// TIA Portal project "Lagerbereich_0" (V20)

(* hardware
DEVICE "S7-1500/ET200MP-Station_1"  S7-1500 station
   slot 0: "Profilschiene_0"  Rack  6ES7 590-1***0-0AA0
   slot 1: "PLC_1"  CPU 1513-1 PN  6ES7 513-1AM03-0AB0  V4.0
      slot 3: "CPU-Display_1"  6ES7591-1AA00-0AA0
      slot 32768: "PROFINET-Schnittstelle_1"  X1
         slot 32769: "Port_1"  X1 P1
         slot 32770: "Port_2"  X1 P2
      slot 34817: "Virtual CP interface port_1"  Virtual CP interface port  Virtual CP interface port FW V4.0
   slot 2: "DI 16x24VDC BA_1"  DI 16x24VDC BA  6ES7 521-1BH10-0AA0  V1.1
   slot 3: "DQ 16x24VDC/0.5A ST_1"  DQ 16x24VDC/0.5A ST  6ES7 522-1BH00-0AB0  V2.0
   slot 4: "AI 8xU/I/R/RTD BA_2"  AI 8xU/I/R/RTD BA  6ES7 531-7QF00-0AB0  V1.0
   slot 5: "AQ 8xU/I HS_2"  AQ 8xU/I HS  6ES7 532-5HF00-0AB0  V2.2
DEVICE "HMI_1"  TP700 Comfort
   slot 0: "HMI_1"  TP700 Comfort  6AV2 124-0GC01-0AX0  17.0.0.0
   slot 1: "HMI_RT_1"  TP700 Comfort  6AV2 124-0GC01-0AX0  17.0.0.0
   slot 5: "HMI_1.IE_CP_1"  PROFINET Interface  17.0.0.0
      slot 1: "PROFINET Schnittstelle_1"  PROFINET Interface
         slot 1: "Port_1"  Port
         slot 2: "Port_2"  Port
   slot 7: "HMI_1.MPI/DP_CP_1"  MPI/DP Interface  17.0.0.0
*)

// ===== PLC "PLC_1"  CPU 1513-1 PN =====

VAR_GLOBAL   // PLC tag table "Eingaenge"
   "1B1" AT %E0.0 : Bool;   // Lichttaster Eingang (LS1)
   "2B1" AT %E0.1 : Bool;   // Lichttaster Ausgang (LS2)
END_VAR

VAR_GLOBAL   // PLC tag table "Ausgaenge"
   "H1" AT %A0.0 : Bool;   // Leuchte leer (P1)
   "H2" AT %A0.1 : Bool;   // Leuchte 10-40% (P2)
   "H3" AT %A0.2 : Bool;   // Leuchte 50% (P3)
   "H4" AT %A0.3 : Bool;   // Leuchte 60-90% (P4)
   "H5" AT %A0.4 : Bool;   // Leuchte voll (P5)
   "1M1" AT %A0.5 : Bool;   // Schranke
   "D1" AT %AD30 : UDInt;   // Display Anzeige Pakete
   "2M1" AT %A1.0 : Bool;   // Band 1
   "2M2" AT %A1.1 : Bool;   // Band 2
   "2M3" AT %A1.2 : Bool;   // Band 3
   "2M4" AT %A1.3 : Bool;   // Band 4
   "2M5" AT %A1.4 : Bool;   // Band 5
   "2M6" AT %A1.5 : Bool;   // Band 6
   "2M7" AT %A1.6 : Bool;   // Band 7
   "2M8" AT %A1.7 : Bool;   // Band 8
END_VAR

DATA_BLOCK "HMI_Schnittstelle"   // DB100
{ S7_Optimized_Access := 'TRUE' }
VERSION : 0.1
   VAR
      Eingaenge : Struct
         "1B1" : Bool;   // Lichttaster Eingang (LS1)
         "2B1" : Bool;   // Lichttaster Ausgang (LS2)
      END_STRUCT;
      Ausgaenge : Struct
         H1 : Bool;   // Leuchte leer (P1)
         H2 : Bool;   // Leuchte 10-40% (P2)
         H3 : Bool;   // Leuchte 50% (P3)
         H4 : Bool;   // Leuchte 60-90% (P4)
         H5 : Bool;   // Leuchte voll (P5)
         "1M1" : Bool;   // Schranke
         Baender : Bool;
         D1 : UDInt;   // Display Anzeige Pakete
         "2M1" : Bool;   // Band 1
         "2M2" : Bool;   // Band 2
         "2M3" : Bool;   // Band 3
         "2M4" : Bool;   // Band 4
         "2M5" : Bool;   // Band 5
         "2M6" : Bool;   // Band 6
         "2M7" : Bool;   // Band 7
         "2M8" : Bool;   // Band 8
      END_STRUCT;
      Betriebsart : Struct
         Hand : Bool := TRUE;
         Automatik : Bool;
      END_STRUCT;
      Lagerbereich : Struct
         Lagerplatz : Array[0..9] of Bool;
      END_STRUCT;
      "CASE" : Bool;
      btnCase : Bool;
   END_VAR
BEGIN
END_DATA_BLOCK

// folder: Anlagensteuerung

DATA_BLOCK "IDB_Anlage"   // DB1
{ S7_Optimized_Access := 'TRUE' }
VERSION : 0.1
// stored: InstanceOfName Ein_Anlage
"Ein_Anlage"
BEGIN
END_DATA_BLOCK

// folder: Logik

DATA_BLOCK "IDB_Schrankensteuerung"   // DB2
{ S7_Optimized_Access := 'TRUE' }
VERSION : 0.1
// stored: InstanceOfName Schrankensteuerung
"Schrankensteuerung"
BEGIN
END_DATA_BLOCK

DATA_BLOCK "IDB_Leuchtensteuerung_IF"   // DB10
{ S7_Optimized_Access := 'TRUE' }
VERSION : 0.1
// stored: InstanceOfName Prog_Steuerung_IF
"Prog_Steuerung_IF"
BEGIN
END_DATA_BLOCK

DATA_BLOCK "IDB_Leuchtensteuerung_CASE"   // DB20
{ S7_Optimized_Access := 'TRUE' }
VERSION : 0.1
// stored: InstanceOfName Prog_Steuerung_CASE
"Prog_Steuerung_CASE"
BEGIN
END_DATA_BLOCK

// folder: (top level)

ORGANIZATION_BLOCK "Main"   // OB1, FBD, ProgramCycle
TITLE = "Main Program Sweep (Cycle)"
{ S7_Optimized_Access := 'TRUE' }
VERSION : 0.1
   VAR_INPUT
      Initial_Call : Bool;   // Initial call of this OB
      Remanence : Bool;   // =True, if remanent data are available
   END_VAR
BEGIN

REGION Network 1: Lichttaster Eingang (LS1)
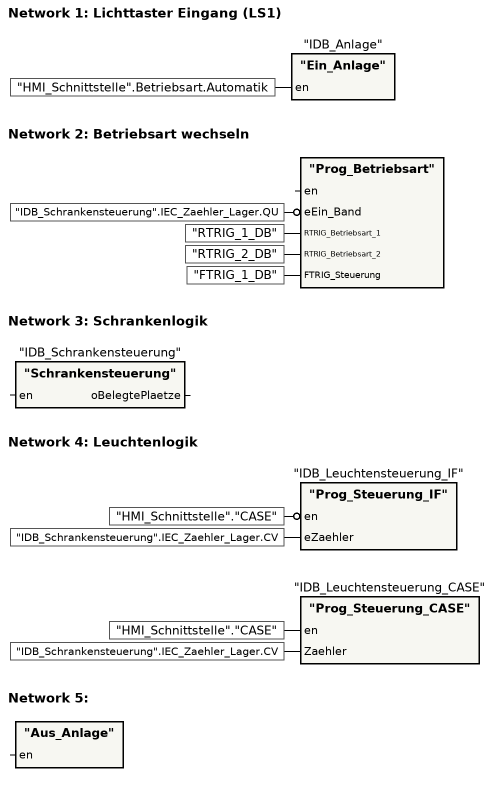
   IF "HMI_Schnittstelle".Betriebsart.Automatik THEN
       "IDB_Anlage"();   // "Ein_Anlage"
   END_IF;
END_REGION

REGION Network 2: Betriebsart wechseln
   "Prog_Betriebsart"(eEin_Band := NOT "IDB_Schrankensteuerung".IEC_Zaehler_Lager.QU,
                      RTRIG_Betriebsart_1 := "RTRIG_1_DB",
                      RTRIG_Betriebsart_2 := "RTRIG_2_DB",
                      FTRIG_Steuerung := "FTRIG_1_DB");
END_REGION

REGION Network 3: Schrankenlogik
   "IDB_Schrankensteuerung"();   // "Schrankensteuerung"
END_REGION

REGION Network 4: Leuchtenlogik
   IF NOT "HMI_Schnittstelle"."CASE" THEN
       "IDB_Leuchtensteuerung_IF"(eZaehler := "IDB_Schrankensteuerung".IEC_Zaehler_Lager.CV);   // "Prog_Steuerung_IF"
   END_IF;
   IF "HMI_Schnittstelle"."CASE" THEN
       "IDB_Leuchtensteuerung_CASE"(Zaehler := "IDB_Schrankensteuerung".IEC_Zaehler_Lager.CV);   // "Prog_Steuerung_CASE"
   END_IF;
END_REGION

REGION Network 5
   "Aus_Anlage"();
END_REGION
END_ORGANIZATION_BLOCK

// folder: Anlagensteuerung

FUNCTION_BLOCK "Ein_Anlage"   // FB1, FBD
{ S7_Optimized_Access := 'TRUE' }
VERSION : 0.1
BEGIN

REGION Network 1 (SCL): Sensoren
   "HMI_Schnittstelle".Eingaenge."1B1" := NOT "1B1";
   "HMI_Schnittstelle".Eingaenge."2B1" := NOT "2B1";
END_REGION
END_FUNCTION_BLOCK

FUNCTION "Aus_Anlage" : Void   // FC1, FBD
{ S7_Optimized_Access := 'TRUE' }
VERSION : 0.1
BEGIN

REGION Network 1 (SCL): Band 1
   "2M1" := "HMI_Schnittstelle".Ausgaenge."2M1";
   "2M2" := "HMI_Schnittstelle".Ausgaenge."2M2";
   "2M3" := "HMI_Schnittstelle".Ausgaenge."2M3";
   "2M4" := "HMI_Schnittstelle".Ausgaenge."2M4";
   "2M5" := "HMI_Schnittstelle".Ausgaenge."2M5";
   "2M6" := "HMI_Schnittstelle".Ausgaenge."2M6";
   "2M7" := "HMI_Schnittstelle".Ausgaenge."2M7";
   "2M8" := "HMI_Schnittstelle".Ausgaenge."2M8";
END_REGION

REGION Network 2 (SCL): Leuchten
   "H1" := "HMI_Schnittstelle".Ausgaenge.H1;
   "H2" := "HMI_Schnittstelle".Ausgaenge.H2;
   "H3" := "HMI_Schnittstelle".Ausgaenge.H3;
   "H4" := "HMI_Schnittstelle".Ausgaenge.H4;
   "H5" := "HMI_Schnittstelle".Ausgaenge.H5;
END_REGION

REGION Network 3 (SCL): Schranke
   "1M1" := "HMI_Schnittstelle".Ausgaenge."1M1";
END_REGION

REGION Network 4 (SCL): Display
   "D1" := "HMI_Schnittstelle".Ausgaenge.D1;
END_REGION
END_FUNCTION

// folder: Logik

FUNCTION_BLOCK "Schrankensteuerung"   // FB2, FBD
{ S7_Optimized_Access := 'TRUE' }
VERSION : 0.1
   VAR_OUTPUT
      oBelegtePlaetze : Int;
   END_VAR
   VAR
      FTRIG_MDB_1B1 : F_TRIG;
      FTRIG_MDB_2B1 : F_TRIG;
   END_VAR
   VAR RETAIN
      IEC_Zaehler_Lager : CTUD_INT;
   END_VAR
   VAR CONSTANT
      cGesamtPlaetze : Int := 10;
   END_VAR
BEGIN

REGION Network 1 (SCL): Flanken Lichttaster
   #FTRIG_MDB_1B1(CLK:= "HMI_Schnittstelle".Eingaenge."1B1");
   #FTRIG_MDB_2B1(CLK:= "HMI_Schnittstelle".Eingaenge."2B1");
END_REGION

REGION Network 2 (SCL): Zählersteuerung
   #IEC_Zaehler_Lager(CU := #FTRIG_MDB_1B1.Q AND #oBelegtePlaetze < #cGesamtPlaetze,
                      CD := #FTRIG_MDB_2B1.Q AND #oBelegtePlaetze > 0,
                      PV := #cGesamtPlaetze,
                      CV=> #oBelegtePlaetze);

   "HMI_Schnittstelle".Ausgaenge.D1 := INT_TO_UDINT(#oBelegtePlaetze);
END_REGION

REGION Network 3 (SCL): Schrankensteuerung
   "HMI_Schnittstelle".Ausgaenge."1M1" := #IEC_Zaehler_Lager.QU;
END_REGION
END_FUNCTION_BLOCK

FUNCTION_BLOCK "Prog_Steuerung_IF"   // FB10, FBD
{ S7_Optimized_Access := 'TRUE' }
VERSION : 0.1
   VAR_INPUT
      eZaehler : UDInt;
   END_VAR
   VAR
      Prozentwert : UInt;
   END_VAR
   VAR CONSTANT
      cGesamtPlaetze : Int := 10;
   END_VAR
BEGIN

REGION Network 1 (SCL): Leuchtensteuerung
   // Wandle den Zähler in einen Prozentwert um
   #Prozentwert := REAL_TO_UINT((UDINT_TO_REAL(#eZaehler) / #cGesamtPlaetze) * 100);


   // Eingänge zurücksetzen
   "HMI_Schnittstelle".Ausgaenge.H1 := FALSE;
   "HMI_Schnittstelle".Ausgaenge.H2 := FALSE;
   "HMI_Schnittstelle".Ausgaenge.H3 := FALSE;
   "HMI_Schnittstelle".Ausgaenge.H4 := FALSE;
   "HMI_Schnittstelle".Ausgaenge.H5 := FALSE;


   IF #Prozentwert < 10 THEN
       "HMI_Schnittstelle".Ausgaenge.H1 := TRUE;
   ELSIF #Prozentwert >= 10 AND #Prozentwert < 50 THEN
       "HMI_Schnittstelle".Ausgaenge.H2 := TRUE;
   ELSIF #Prozentwert = 50 THEN
       "HMI_Schnittstelle".Ausgaenge.H3 := TRUE;
   ELSIF #Prozentwert > 50 AND #Prozentwert <= 90 THEN
       "HMI_Schnittstelle".Ausgaenge.H4 := TRUE;
   ELSIF #Prozentwert > 90 THEN
       "HMI_Schnittstelle".Ausgaenge.H5 := TRUE;
   END_IF;
END_REGION
END_FUNCTION_BLOCK

FUNCTION_BLOCK "Prog_Steuerung_CASE"   // FB20, FBD
{ S7_Optimized_Access := 'TRUE' }
VERSION : 0.1
   VAR_INPUT
      Zaehler : UDInt;
   END_VAR
   VAR
      Prozentwert : UInt;
   END_VAR
   VAR CONSTANT
      cGesamtPlaetze : Int := 10;
   END_VAR
BEGIN

REGION Network 1 (SCL): Leuchtensteuerung
   // Wandle den Zähler in einen Prozentwert um
   #Prozentwert := REAL_TO_UINT((UDINT_TO_REAL(#Zaehler) / #cGesamtPlaetze) * 100);


   // Eingänge zurücksetzen
   "HMI_Schnittstelle".Ausgaenge.H1 := FALSE;
   "HMI_Schnittstelle".Ausgaenge.H2 := FALSE;
   "HMI_Schnittstelle".Ausgaenge.H3 := FALSE;
   "HMI_Schnittstelle".Ausgaenge.H4 := FALSE;
   "HMI_Schnittstelle".Ausgaenge.H5 := FALSE;

   CASE #Prozentwert OF
       0..9:// < 10
           "HMI_Schnittstelle".Ausgaenge.H1 := TRUE;
       10..49:// >= 10 AND < 50
           "HMI_Schnittstelle".Ausgaenge.H2 := TRUE;
       50:// = 50
           "HMI_Schnittstelle".Ausgaenge.H3 := TRUE;
       51..90:// > 50 AND <= 90
           "HMI_Schnittstelle".Ausgaenge.H4 := TRUE;
       91..100:// > 90
           "HMI_Schnittstelle".Ausgaenge.H5 := TRUE;
       ELSE;
   END_CASE;
END_REGION
END_FUNCTION_BLOCK

FUNCTION "Prog_Betriebsart" : Void   // FC2, FBD
{ S7_Optimized_Access := 'TRUE' }
VERSION : 0.1
   VAR_INPUT
      eEin_Band : Bool;
   END_VAR
   VAR_IN_OUT
      RTRIG_Betriebsart_1 : R_TRIG;
      RTRIG_Betriebsart_2 : R_TRIG;
      FTRIG_Steuerung : F_TRIG;
   END_VAR
   VAR_TEMP
      tmpCase : Bool;
   END_VAR
BEGIN

REGION Network 1 (SCL)
   #RTRIG_Betriebsart_1(CLK := "HMI_Schnittstelle".Betriebsart.Hand);
   #RTRIG_Betriebsart_2(CLK := "HMI_Schnittstelle".Betriebsart.Automatik);

   "HMI_Schnittstelle".Betriebsart.Automatik := #RTRIG_Betriebsart_1.Q XOR "HMI_Schnittstelle".Betriebsart.Automatik;
   "HMI_Schnittstelle".Betriebsart.Hand := #RTRIG_Betriebsart_2.Q XOR "HMI_Schnittstelle".Betriebsart.Hand;
END_REGION

REGION Network 2 (SCL)
   #FTRIG_Steuerung(CLK:= "HMI_Schnittstelle".btnCase);

   IF #FTRIG_Steuerung.Q THEN
       "HMI_Schnittstelle"."CASE" := NOT "HMI_Schnittstelle"."CASE";
   END_IF;
END_REGION

REGION Network 3 (SCL): Bandsteuerung
   "HMI_Schnittstelle".Ausgaenge.Baender := "HMI_Schnittstelle".Betriebsart.Automatik;

   "HMI_Schnittstelle".Ausgaenge."2M1" := #eEin_Band;
   "HMI_Schnittstelle".Ausgaenge."2M2" := "HMI_Schnittstelle".Ausgaenge.Baender;
   "HMI_Schnittstelle".Ausgaenge."2M3" := "HMI_Schnittstelle".Ausgaenge.Baender;
   "HMI_Schnittstelle".Ausgaenge."2M4" := "HMI_Schnittstelle".Ausgaenge.Baender;
   "HMI_Schnittstelle".Ausgaenge."2M5" := "HMI_Schnittstelle".Ausgaenge.Baender;
   "HMI_Schnittstelle".Ausgaenge."2M6" := "HMI_Schnittstelle".Ausgaenge.Baender;
   "HMI_Schnittstelle".Ausgaenge."2M7" := "HMI_Schnittstelle".Ausgaenge.Baender;
   "HMI_Schnittstelle".Ausgaenge."2M8" := "HMI_Schnittstelle".Ausgaenge.Baender;
END_REGION
END_FUNCTION

// ===== library types =====

// folder: LGF/0 Bit logic operations

FUNCTION "LGF_BitToggle" : DWord   // FC10033, SCL
TITLE = LGF_BitToggle
{ S7_Optimized_Access := 'TRUE' }
AUTHOR : Siemens_SIMATIC_Systems_Support
FAMILY : LGF
NAME : LGF_BitToggle
// Dieser Baustein toggelt (von TRUE nach FALSE und umgekehrt) ein Bit an vorgegebener Stelle in einer Variablen vom Datentyp DWORD.    
// Anstelle von DWord kann auch Word und Byte verwendet werden, indem der übergebene Parameter mit z. B. BYTE_TO_DWORD und das Ergebnis mit DWORD_TO_BYTE konvertiert wird.
// This block toggles (from TRUE to FALSE and vice versa) a bit at a predefined position in a variable of the data type DWORD.  
// Alternatively, Word and Byte can be used instead of DWord by converting the passed parameter with, for example, BYTE_TO_DWORD and the result with DWORD_TO_BYTE
   VAR_INPUT
      value : DWord;   // Tag where the bit has to be toggled / Variable, an der das Bit getoggelt wird.
      bitNo : USInt;   // Bit number to be toggled in the “value” parameter. / Bitnummer, die im Parameter "value" getoggelt werden soll.
   END_VAR
   // Ret_Val : Tag with toggled bit / Variable mit getoggeltem Bit.
   VAR CONSTANT
      TRUE_BOOL_BIT : DWord := 16#0001;   // Just one bit which is true, to shift in Dword for masking / Ein einzelnes Bit mit Wert := TRUE zum schieben im Dword und zur Maskierung
      MAX_NO_OF_BITS : USInt := 32;   // Maximum bits in a DWord = 32 / Maximalanzahl an Bits in einem Dword = 32
   END_VAR
BEGIN
   REGION BLOCK INFO HEADER
     //===============================================================================
     // SIEMENS AG / (c)Copyright 2019
     //-------------------------------------------------------------------------------
     // Title:            LGF_BitToggle
     // Comment/Function: Toggle bit in elementary datatype - DWord
     //                   can be used for Word and Byte as well, by convert
     //                   the passed paramter and the result using for e.g. Dword_to_Byte
     // Library/Family:   LGF (Library General Functions)
     // Author:           Siemens Digital Industry
     // Tested with:      CPU1212C DC/DC/DC FW:V4.2
     // Engineering:      TIA Portal V15.1
     // Restrictions:     ENO not in use, set to true, no error handling
     // Requirements:     PLC (S7-1200 / S7-1500)
     //-------------------------------------------------------------------------------
     // Change log table:
     // Version  | Date       | Expert in charge         | Changes applied
     // 01.00.00 | 06.06.2015 | Siemens Industry Support | first release
     // 03.00.00 | 23.04.2020 | Siemens Industry Support | Set version to V3.0.0
     //                         harmonize the version of the whole library
     // 03.00.01 | 19.01.2021 | Simatic Systems Support
     //                         Insert documentation
     //===============================================================================
   END_REGION

   REGION Logic
     // toggle the bit in tag
     // shift one true bit into given position
     // concatenate value then with XOR resets the bit on the given position
     #LGF_BitToggle := #value XOR SHL(IN := #TRUE_BOOL_BIT, N := (#bitNo MOD #MAX_NO_OF_BITS));

     // no error handling needed
     ENO := TRUE;
   END_REGION
END_FUNCTION

(* ===== HMI "HMI_RT_1" =====
system functions are stored by id; their names below are inferred from use
connection "HMI_Verbindung_1": ETHERNET, S7_1500_OMS

HMI tags "Standard-Variablentabelle"
   "HMI_Schnittstelle_Eingaenge_1B1" : Bool = PLC HMI_Schnittstelle.Eingaenge.1B1, 100 ms
   "HMI_Schnittstelle_Eingaenge_2B1" : Bool = PLC HMI_Schnittstelle.Eingaenge.2B1, 100 ms
   "HMI_Schnittstelle_Ausgaenge_1M1" : Bool = PLC HMI_Schnittstelle.Ausgaenge.1M1, 100 ms
   "HMI_Schnittstelle_Ausgaenge_D1" : UDInt = PLC HMI_Schnittstelle.Ausgaenge.D1, 100 ms
   "HMI_Schnittstelle_Ausgaenge_H3" : Bool = PLC HMI_Schnittstelle.Ausgaenge.H3, 500 ms
   "HMI_Schnittstelle_Ausgaenge_H4" : Bool = PLC HMI_Schnittstelle.Ausgaenge.H4, 500 ms
   "HMI_Schnittstelle_Ausgaenge_H2" : Bool = PLC HMI_Schnittstelle.Ausgaenge.H2, 500 ms
   "HMI_Schnittstelle_Ausgaenge_H1" : Bool = PLC HMI_Schnittstelle.Ausgaenge.H1, 500 ms
   "HMI_Schnittstelle_Ausgaenge_H5" : Bool = PLC HMI_Schnittstelle.Ausgaenge.H5, 500 ms
   "HMI_Schnittstelle_Betriebsart_Hand" : Bool = PLC HMI_Schnittstelle.Betriebsart.Hand, 100 ms
   "HMI_Schnittstelle_Betriebsart_Automatik" : Bool = PLC HMI_Schnittstelle.Betriebsart.Automatik, 100 ms
   "HMI_Schnittstelle_CASE" : Bool = PLC HMI_Schnittstelle.CASE, 100 ms
   "HMI_Schnittstelle_btnCase" : Bool = PLC HMI_Schnittstelle.btnCase, 100 ms

screen "01_Startseite" 800x480
   Rectangle "Rechteck_1" at 25,140 size 10x200
      Appearance <- "HMI_Schnittstelle_Ausgaenge_1M1"
   IOField "EA-Feld_1" at 352,224 size 96x32; FormatPattern 99
      ProcessValue <- "HMI_Schnittstelle_Ausgaenge_D1"
   Circle "Kreis_1" at 384,100 size 32x32
      Appearance <- "HMI_Schnittstelle_Ausgaenge_H3"
   Circle "Kreis_2" at 344,100 size 32x32
      Appearance <- "HMI_Schnittstelle_Ausgaenge_H2"
   Circle "Kreis_3" at 424,100 size 32x32
      Appearance <- "HMI_Schnittstelle_Ausgaenge_H4"
   Circle "Kreis_4" at 304,100 size 32x32
      Appearance <- "HMI_Schnittstelle_Ausgaenge_H1"
   Circle "Kreis_5" at 464,100 size 32x32
      Appearance <- "HMI_Schnittstelle_Ausgaenge_H5"
   Button "Schaltfläche_3" at 304,348 size 96x32; TextOff 'Hand'
      Appearance <- "HMI_Schnittstelle_Betriebsart_Hand"
      on Press: SetBit("HMI_Schnittstelle_Betriebsart_Hand")
   Button "Schaltfläche_4" at 400,348 size 96x32; TextOff 'Auto'
      Appearance <- "HMI_Schnittstelle_Betriebsart_Automatik"
      on Press: SetBit("HMI_Schnittstelle_Betriebsart_Automatik")
   Button "Schaltfläche_5" at 352,390 size 96x32; TextOff 'CASE'
      Appearance <- "HMI_Schnittstelle_CASE"
      on Press: function_b14e0dd5("HMI_Schnittstelle_btnCase", 0)
   Button "Schaltfläche_7" at 652,224 size 48x32; TextOff '2B1'
      Appearance <- "HMI_Schnittstelle_Eingaenge_2B1"
      on Press: function_b14e0dd5("HMI_Schnittstelle_Eingaenge_2B1", 0)
      Visibility <- "HMI_Schnittstelle_Betriebsart_Automatik"
   Button "Schaltfläche_6" at 100,224 size 48x32; TextOff '1B1'
      Appearance <- "HMI_Schnittstelle_Eingaenge_1B1"
      on Press: function_b14e0dd5("HMI_Schnittstelle_Eingaenge_1B1", 0)
      Visibility <- "HMI_Schnittstelle_Betriebsart_Automatik"
   Rectangle "Rechteck_4" at 100,224 size 48x32
      Appearance <- "HMI_Schnittstelle_Eingaenge_1B1"
      Visibility <- "HMI_Schnittstelle_Betriebsart_Hand"
   TextField "Textfeld_1" at 100,224 size 48x32; Text '1B1'
   Rectangle "Rechteck_5" at 652,224 size 48x32
      Visibility <- "HMI_Schnittstelle_Betriebsart_Hand"
      Appearance <- "HMI_Schnittstelle_Eingaenge_2B1"
   TextField "Textfeld_2" at 652,224 size 48x32; Text '2B1'
   Group "Group" at 100,224 size 48x32
   Group "Group_1" at 652,224 size 48x32
*)